// TIA Portal project "HEAT-1-CADIZ-V24" (V20) (continued)

       CASE #modeRequest OF
           1: // ======= Conceder control a KukaControl =========
               // Requisito: que el otro lado (Supervisor) esté ocioso (Queda por ajustar)
               IF #safeAllOk AND (NOT #autoBusy) THEN

                   // 1) Fijar modo efectivo → AutoExtSeq cargará PGNO = 1
                   #modeEffective := USINT#1;

                   // 2) Aún no estamos listos hasta que AutoExtSeq termine
                   "PlcStatus".mode.ready := FALSE;

                   // 3) Señal PNIO al robot para que salga del bucle autoloop.src (CASE 1 del cell.src)
                   #enterCellCase1 := TRUE;

                   // 4) Arranque de AutoExt: PULSO 1-scan a %M770.0
                   #startAutoExt := TRUE;

                   // 5) Handshake a la HMI con el MISMO seq que se recibió
                   "PlcStatus".exec.ackSeq := #modeReqSeq;
                   "PlcStatus".exec.accepted := TRUE;  // 1 scan
                   "PlcStatus".exec.done := TRUE;  // 1 scan
               END_IF;

           2: // ======= Conceder control a Supervisor/VisualScan =========
               // Requisito: que KukaControl esté ocioso
               IF #safeAllOk AND (NOT #servBusy) THEN

                   // 1) Fijar modo efectivo → AutoExtSeq cargará PGNO = 2
                   #modeEffective := USINT#2;

                   // 2) Aún no estamos listos hasta que AutoExtSeq termine
                   "PlcStatus".mode.ready := FALSE;

                   // 3) Señal PNIO al robot para que salga del bucle actual autoloopsup.src (CASE 2 del cell.src)
                   #enterCellCase2 := TRUE;

                   // 4) Arranque de AutoExt: PULSO 1-scan a %M770.0
                   #startAutoExt := TRUE;

                   // 5) Handshake a la HMI
                   "PlcStatus".exec.ackSeq := #modeReqSeq;
                   "PlcStatus".exec.accepted := TRUE;
                   "PlcStatus".exec.done := TRUE;
               END_IF;
       END_CASE;

   END_IF;
END_REGION
END_FUNCTION_BLOCK

FUNCTION_BLOCK "KukaControlSeq"   // FB21, LAD
{ S7_Optimized_Access := 'TRUE' }
VERSION : 0.1
   VAR
      rEnterAuto : R_TRIG;
   END_VAR
   VAR_TEMP
      _clear990 : Bool;
   END_VAR
BEGIN

REGION Network 2: Envia posiciones a la aplicacion KukaControl
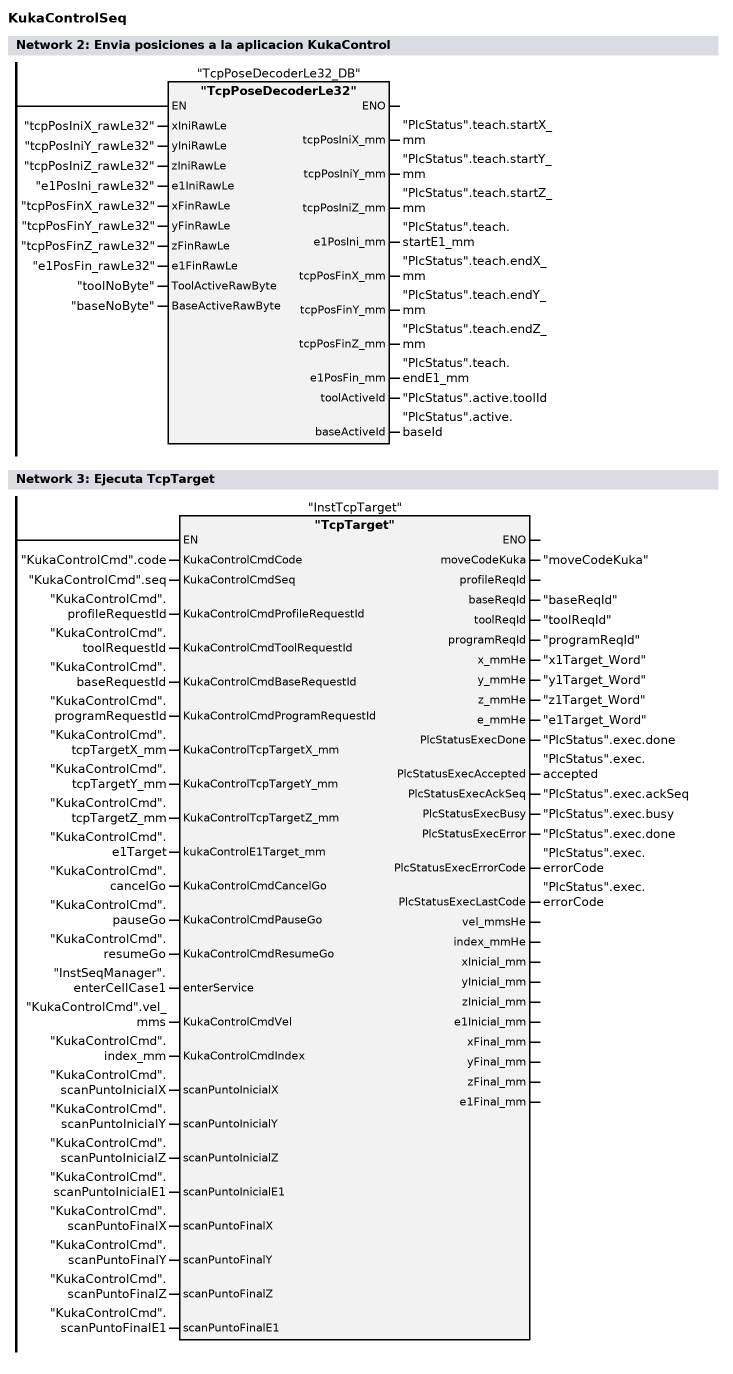
   RUNG wire#powerrail
      "TcpPoseDecoderLe32_DB"(xIniRawLe := "tcpPosIniX_rawLe32", yIniRawLe := "tcpPosIniY_rawLe32", zIniRawLe := "tcpPosIniZ_rawLe32", e1IniRawLe := "e1PosIni_rawLe32", xFinRawLe := "tcpPosFinX_rawLe32", yFinRawLe := "tcpPosFinY_rawLe32", zFinRawLe := "tcpPosFinZ_rawLe32", e1FinRawLe := "e1PosFin_rawLe32", ToolActiveRawByte := "toolNoByte", BaseActiveRawByte := "baseNoByte", tcpPosIniX_mm => "PlcStatus".teach.startX_mm, tcpPosIniY_mm => "PlcStatus".teach.startY_mm, tcpPosIniZ_mm => "PlcStatus".teach.startZ_mm, e1PosIni_mm => "PlcStatus".teach.startE1_mm, tcpPosFinX_mm => "PlcStatus".teach.endX_mm, tcpPosFinY_mm => "PlcStatus".teach.endY_mm, tcpPosFinZ_mm => "PlcStatus".teach.endZ_mm, e1PosFin_mm => "PlcStatus".teach.endE1_mm, toolActiveId => "PlcStatus".active.toolId, baseActiveId => "PlcStatus".active.baseId)
   END_RUNG
   // the same network as SCL:
   "TcpPoseDecoderLe32_DB"(xIniRawLe := "tcpPosIniX_rawLe32",   // "TcpPoseDecoderLe32"
                           yIniRawLe := "tcpPosIniY_rawLe32",
                           zIniRawLe := "tcpPosIniZ_rawLe32",
                           e1IniRawLe := "e1PosIni_rawLe32",
                           xFinRawLe := "tcpPosFinX_rawLe32",
                           yFinRawLe := "tcpPosFinY_rawLe32",
                           zFinRawLe := "tcpPosFinZ_rawLe32",
                           e1FinRawLe := "e1PosFin_rawLe32",
                           ToolActiveRawByte := "toolNoByte",
                           BaseActiveRawByte := "baseNoByte",
                           tcpPosIniX_mm => "PlcStatus".teach.startX_mm,
                           tcpPosIniY_mm => "PlcStatus".teach.startY_mm,
                           tcpPosIniZ_mm => "PlcStatus".teach.startZ_mm,
                           e1PosIni_mm => "PlcStatus".teach.startE1_mm,
                           tcpPosFinX_mm => "PlcStatus".teach.endX_mm,
                           tcpPosFinY_mm => "PlcStatus".teach.endY_mm,
                           tcpPosFinZ_mm => "PlcStatus".teach.endZ_mm,
                           e1PosFin_mm => "PlcStatus".teach.endE1_mm,
                           toolActiveId => "PlcStatus".active.toolId,
                           baseActiveId => "PlcStatus".active.baseId);
END_REGION

REGION Network 3: Ejecuta TcpTarget
   RUNG wire#powerrail
      "InstTcpTarget"(KukaControlCmdCode := "KukaControlCmd".code, KukaControlCmdSeq := "KukaControlCmd".seq, KukaControlCmdProfileRequestId := "KukaControlCmd".profileRequestId, KukaControlCmdToolRequestId := "KukaControlCmd".toolRequestId, KukaControlCmdBaseRequestId := "KukaControlCmd".baseRequestId, KukaControlCmdProgramRequestId := "KukaControlCmd".programRequestId, KukaControlTcpTargetX_mm := "KukaControlCmd".tcpTargetX_mm, KukaControlTcpTargetY_mm := "KukaControlCmd".tcpTargetY_mm, KukaControlTcpTargetZ_mm := "KukaControlCmd".tcpTargetZ_mm, kukaControlE1Target_mm := "KukaControlCmd".e1Target, KukaControlCmdCancelGo := "KukaControlCmd".cancelGo, KukaControlCmdPauseGo := "KukaControlCmd".pauseGo, KukaControlCmdResumeGo := "KukaControlCmd".resumeGo, enterService := "InstSeqManager".enterCellCase1, KukaControlCmdVel := "KukaControlCmd".vel_mms, KukaControlCmdIndex := "KukaControlCmd".index_mm, scanPuntoInicialX := "KukaControlCmd".scanPuntoInicialX, scanPuntoInicialY := "KukaControlCmd".scanPuntoInicialY, scanPuntoInicialZ := "KukaControlCmd".scanPuntoInicialZ, scanPuntoInicialE1 := "KukaControlCmd".scanPuntoInicialE1, scanPuntoFinalX := "KukaControlCmd".scanPuntoFinalX, scanPuntoFinalY := "KukaControlCmd".scanPuntoFinalY, scanPuntoFinalZ := "KukaControlCmd".scanPuntoFinalZ, scanPuntoFinalE1 := "KukaControlCmd".scanPuntoFinalE1, moveCodeKuka => "moveCodeKuka", profileReqId =>, baseReqId => "baseReqId", toolReqId => "toolReqId", programReqId => "programReqId", x_mmHe => "x1Target_Word", y_mmHe => "y1Target_Word", z_mmHe => "z1Target_Word", e_mmHe => "e1Target_Word", PlcStatusExecDone => "PlcStatus".exec.done, PlcStatusExecAccepted => "PlcStatus".exec.accepted, PlcStatusExecAckSeq => "PlcStatus".exec.ackSeq, PlcStatusExecBusy => "PlcStatus".exec.busy, PlcStatusExecError => "PlcStatus".exec.done, PlcStatusExecErrorCode => "PlcStatus".exec.errorCode, PlcStatusExecLastCode => "PlcStatus".exec.errorCode, vel_mmsHe =>, index_mmHe =>, xInicial_mm =>, yInicial_mm =>, zInicial_mm =>, e1Inicial_mm =>, xFinal_mm =>, yFinal_mm =>, zFinal_mm =>, e1Final_mm =>)
   END_RUNG
   // the same network as SCL:
   "InstTcpTarget"(KukaControlCmdCode := "KukaControlCmd".code,   // "TcpTarget"
                   KukaControlCmdSeq := "KukaControlCmd".seq,
                   KukaControlCmdProfileRequestId := "KukaControlCmd".profileRequestId,
                   KukaControlCmdToolRequestId := "KukaControlCmd".toolRequestId,
                   KukaControlCmdBaseRequestId := "KukaControlCmd".baseRequestId,
                   KukaControlCmdProgramRequestId := "KukaControlCmd".programRequestId,
                   KukaControlTcpTargetX_mm := "KukaControlCmd".tcpTargetX_mm,
                   KukaControlTcpTargetY_mm := "KukaControlCmd".tcpTargetY_mm,
                   KukaControlTcpTargetZ_mm := "KukaControlCmd".tcpTargetZ_mm,
                   kukaControlE1Target_mm := "KukaControlCmd".e1Target,
                   KukaControlCmdCancelGo := "KukaControlCmd".cancelGo,
                   KukaControlCmdPauseGo := "KukaControlCmd".pauseGo,
                   KukaControlCmdResumeGo := "KukaControlCmd".resumeGo,
                   enterService := "InstSeqManager".enterCellCase1,
                   KukaControlCmdVel := "KukaControlCmd".vel_mms,
                   KukaControlCmdIndex := "KukaControlCmd".index_mm,
                   scanPuntoInicialX := "KukaControlCmd".scanPuntoInicialX,
                   scanPuntoInicialY := "KukaControlCmd".scanPuntoInicialY,
                   scanPuntoInicialZ := "KukaControlCmd".scanPuntoInicialZ,
                   scanPuntoInicialE1 := "KukaControlCmd".scanPuntoInicialE1,
                   scanPuntoFinalX := "KukaControlCmd".scanPuntoFinalX,
                   scanPuntoFinalY := "KukaControlCmd".scanPuntoFinalY,
                   scanPuntoFinalZ := "KukaControlCmd".scanPuntoFinalZ,
                   scanPuntoFinalE1 := "KukaControlCmd".scanPuntoFinalE1,
                   moveCodeKuka => "moveCodeKuka",
                   baseReqId => "baseReqId",
                   toolReqId => "toolReqId",
                   programReqId => "programReqId",
                   x_mmHe => "x1Target_Word",
                   y_mmHe => "y1Target_Word",
                   z_mmHe => "z1Target_Word",
                   e_mmHe => "e1Target_Word",
                   PlcStatusExecDone => "PlcStatus".exec.done,
                   PlcStatusExecAccepted => "PlcStatus".exec.accepted,
                   PlcStatusExecAckSeq => "PlcStatus".exec.ackSeq,
                   PlcStatusExecBusy => "PlcStatus".exec.busy,
                   PlcStatusExecError => "PlcStatus".exec.done,
                   PlcStatusExecErrorCode => "PlcStatus".exec.errorCode,
                   PlcStatusExecLastCode => "PlcStatus".exec.errorCode);
END_REGION

REGION Network 4 (SCL)
   IF #_clear990 THEN
       "KukaControlCmd".code := 0;                     // no “ensucia” el DB
       #_clear990 := FALSE;
   END_IF;
END_REGION
END_FUNCTION_BLOCK

FUNCTION_BLOCK "SupervisorSeq"   // FB22, LAD
{ S7_Optimized_Access := 'TRUE' }
VERSION : 0.1
   VAR_INPUT
      T_Heartbeat : Time := T#1000ms;   // Periodo del heartbeat PLC
      T_IdCheck : Time := T#2000ms;   // Duración simulada de Identification (comprobaciones)
      enable : Bool;   // Habilita FB -> PLC.plc_ok
      QR_Ready : Bool := true;   // Hay un ID de carrito leído
      CarriageID : String := 'null';   // ID de carrito leído por QR
      TeachAtStart : Bool;   // Teaching (pág. 4): robot en punto de inicio de la siguiente trayectoria
      kukaAtPerspexPos : Bool;   // PA check (Perspex) y Balancing (pág. 6): Robot posicionado en Perspex
      kukaAtGainPos : Bool;   // Gain (pág. 7) -Robot posicionado para Gain
      kukaAtTCGPos : Bool;   // TCG (pág. 8) — multiposición Robot en la posición TCG actual
      kukaAtRefScanStartPos : Bool;   // Robot listo para Scan Ref
      kukaAtInspScanStartPos : Bool;   // Robot listo para Scan Insp
      kukaRefScanFinished : Bool;   // Trayectoria de referencia terminada (robot/UT)
      kukaInspScanFinished : Bool;   // Trayectoria de inspección terminada (robot/UT)
      StartUSReady : Bool := TRUE;   // StartUS (pág. 5): end-effector y precondiciones listas -- True cuando “previous task done”
      MarkingDone : Bool;   // Pre-eval / marcado (pág. 13) -Resultado del marcado (true=OK)
      CmdStopUS : Bool;   // Orden local para Stop US
      CmdBreakUS : Bool;   // Pulso local Break US
      CmdUnbreakUS : Bool;   // Pulso local Unbreak US
   END_VAR
   VAR_OUTPUT
      ActiveStep : Int;   // Espejo local de PLC.step_plc
      AckSourceDbg : Int;   // Código de fuente de ACK (debug local)
      TCG_NextPosReq : Bool;   // PULSO 1 ciclo: mover a la SIGUIENTE posición TCG
      programReqId : Word;
      moveCodeKuka : Word;
      TCG_AdjustMode : Bool;   // LATCH: TRUE mientras estamos en “ajuste TCG”
   END_VAR
   VAR
      tHeartbeat : TON_TIME;
      hbGate : Bool;
      prevStep : Int := -32768;
      firstScan : Bool;
      teachWasRunning : Bool;
      startUSWasRunning : Bool;
      elemWasRunning : Bool;
      balWasRunning : Bool;
      gainWasRunning : Bool;
      scanRefWasRunning : Bool;
      scanInspWasRunning : Bool;
      L_IdEvalDone : Bool;   // // Identification: ya evalué reqId
      L_tcgNext : Bool;
      L_reqRef : Bool;
      L_reqStop : Bool;
      L_reqTcgAdj : Bool;
      L_reqVerif : Bool;
      L_reqPreEval : Bool;
      L_reqIdent : Bool;
      L_reqMark : Bool;
      carriageLatched : Bool;
      validScanParams : Bool;
      waitingNextTCGPos : Bool;
      Cfg_EndEffector : Int;
      Cfg_TeachReq : Bool;
      Cfg_PaCheckReq : Bool;
      Cfg_TcgReq : Bool;
      Cfg_RefName : String;
      PartProgIdx : UInt := 1;   // // index de programa INSP (pieza)
      RefProgIdx : UInt := 1;   // // index de programa REF (pieza)
      tcgIndex : UInt := 1;   // // posición TCG actual
      WantCode : UInt;
      WantProgId : UInt;
      WantToolId : UInt;
      WantIndex : UInt;
      state : Int;
      lastSeq : UInt;
      SupervisorCmdSeq : UInt;
   END_VAR
   VAR_TEMP
      _clear990 : Bool;
      code_int : UInt;
   END_VAR
   VAR CONSTANT
      cSTEP_ID : Int := 1;   // // Pasos (según resumen del PDF, pág. 1)
      cSTEP_TEACH : Int := 2;
      cSTEP_STARTUS : Int := 3;
      cSTEP_PA_BAL : Int := 4;
      cSTEP_GAIN : Int := 5;
      cSTEP_TCG : Int := 6;
      cSTEP_SCAN_REF : Int := 7;
      cSTEP_SCAN_INSP : Int := 8;
      cSTEP_SCAN_REF_VERIF : Int := 9;
      cSTEP_PRE_EVAL : Int := 10;
      cKUKA_REQ_TOOL : UInt := 201;
      cKUKA_GOTO_PERSPEX : UInt := 412;   // mover a Perspex (usa punto enseñado en KRC)
      cKUKA_GOTO_GAIN : UInt := 413;   // mover a Gain
      cKUKA_GOTO_TCG : UInt := 414;   // mover a posición TCG (ARG = index)
      cKUKA_GOTO_REF_START : UInt := 420;   // mover a inicio de Ref (ARG = RefProgIdx)
      cKUKA_GOTO_INSP_START : UInt := 421;   // mover a inicio de Insp (ARG = PartProgIdx)
      cKUKA_RUN_REF_PATH : UInt := 432;   // ejecutar trayectoria de Ref (ARG = RefProgIdx)
      cKUKA_RUN_INSP_PATH : UInt := 433;   // ejecutar trayectoria de Insp (ARG = PartProgIdx)
   END_VAR
BEGIN

REGION Network 1 (SCL)
   // ------------------------------------------------------------------
   // 0) Servicios globales (Heartbeat, housekeeping) — vars generales (pág. 2)
   // ------------------------------------------------------------------
   "PlcStatus".plcOk := #enable;         // espejo de habilitación

   // Heartbeat PLC: toggle con TON (patrón de "compuerta")
   // hbGate se pone TRUE -> TON corre hasta PT -> tHeartbeat.Q = TRUE -> togglamos
   // y bajamos hbGate para reiniciar el ciclo.
   #tHeartbeat(IN := #hbGate,
               PT := #T_Heartbeat);
   IF NOT #hbGate THEN
       #hbGate := TRUE;
   ELSIF #tHeartbeat.Q THEN
       "PlcStatus".heartbeatPlc := NOT "PlcStatus".heartbeatPlc;
       #hbGate := FALSE;
   END_IF;

   // Normalizar paso y espejarlo a salida
   IF ("PlcStatus".stepPlc < #cSTEP_ID) OR ("PlcStatus".stepPlc > #cSTEP_PRE_EVAL) THEN
       "PlcStatus".stepPlc := #cSTEP_ID;
   END_IF;
   #ActiveStep := "PlcStatus".stepPlc;

   // firstScan: 1 ciclo al entrar en cada paso -> útil para resets seguros
   #firstScan := ("PlcStatus".stepPlc <> #prevStep);
   IF #firstScan THEN
       // Limpiamos cualquier "ready/start" que no deba arrastrarse al paso nuevo
       "PlcStatus".startUsReady := FALSE;
       "PlcStatus".stopUsReady := FALSE;
       "PlcStatus".paCheckReady := FALSE;
       "PlcStatus".gainReady := FALSE;
       "PlcStatus".tcgReady := FALSE;
       "PlcStatus".scanRefStart := FALSE;
       "PlcStatus".scanInspStart := FALSE;
       "PlcStatus".markRunning := FALSE;

       // Latches de “estaba corriendo”
       #teachWasRunning := FALSE;
       #startUSWasRunning := FALSE;
       #elemWasRunning := FALSE;
       #balWasRunning := FALSE;
       #gainWasRunning := FALSE;
       #scanRefWasRunning := FALSE;
       #scanInspWasRunning := FALSE;

       // Latches de peticiones (se “arman” al estado actual para evitar disparos al entrar)
       #L_tcgNext := "SupervisorCmd".tcgNextStep;
       #L_reqRef := "SupervisorCmd".reqRefPart;
       #L_reqStop := "SupervisorCmd".reqStopCycle;
       #L_reqTcgAdj := "SupervisorCmd".reqTcgAdj;
       #L_reqVerif := "SupervisorCmd".reqVerif;
       #L_reqPreEval := "SupervisorCmd".reqPreEval;
       #L_reqIdent := "SupervisorCmd".reqIdentificationState;
       #L_reqMark := "SupervisorCmd".reqMark;

       // Identification
       "PlcStatus".idRunning := FALSE;
       #L_IdEvalDone := FALSE;

       // TCG
       #waitingNextTCGPos := ("PlcStatus".stepPlc = #cSTEP_TCG) AND (NOT #kukaAtTCGPos);
       IF "PlcStatus".stepPlc <> #cSTEP_TCG THEN
           #tcgIndex := 1;
       END_IF;

       // Vaciar slot de orden pendiente a robot
       #WantCode := 0;
       #WantProgId := 0;
       #WantToolId := 0;
       #WantIndex := 0;

       #prevStep := "PlcStatus".stepPlc;
   END_IF;

   // ------------------------------------------------------------------
   //[1] MÁQUINA DE ESTADOS (OPC UA + disparos al KUKA por goTrigger)
   // ------------------------------------------------------------------
   CASE "PlcStatus".stepPlc OF

           // ===============================================================
           // 1) IDENTIFICATION (pág. 3)
           // ===============================================================
       #cSTEP_ID:
           // --- Handshake de carriage ID ---
           // FÍSICO: lectura real de QR/PNs/params en KukaControl.
           // El PLC refleja ID leído y valida condiciones base (safety, agua, robot OK).
           // Supervisor.req_carriage_id = TRUE -> el PLC debe mandar:
           //   PLC.carriage_Id (string) y PLC.new_carriage_Id = TRUE
           // Mientras dure la petición. Al bajar la petición, el PLC
           // limpia new_carriage_Id y deja de enviar.
           // req_carriage_id: enviar ID nuevo UNA VEZ mientras Supervisor lo solicite
           IF "SupervisorCmd".reqCarriageId THEN
               IF #QR_Ready AND NOT #carriageLatched  THEN
                   #CarriageID := 'Id de Prueba';
                   "PlcStatus".carriageId := #CarriageID; // escribimos el ID leído
                   "PlcStatus".newCarriageId := TRUE;     // “ID listo”
                   #carriageLatched  := TRUE;              // evita rearmar en el mismo pulso
               END_IF;
           ELSE
               // fin del handshake
               "PlcStatus".newCarriageId := FALSE;
               #carriageLatched  := FALSE;
           END_IF;

           // --- req_id (latch: eval una sola vez en “alto” y decidir salto al bajar) ---
           "PlcStatus".idRunning := "SupervisorCmd".reqId;

           // 1) Primera vez con reqId=TRUE → congelar configuración + calcular id_ok
           IF "SupervisorCmd".reqId AND NOT #L_IdEvalDone THEN
               // Congelar lo que Supervisor ha decidido para el ciclo
               #Cfg_EndEffector := "SupervisorCmd".endEffector;  // 1..5
               #Cfg_TeachReq := "SupervisorCmd".teachReq;
               #Cfg_PaCheckReq := "SupervisorCmd".paCheckReq;
               #Cfg_TcgReq := "SupervisorCmd".tcgReq;
               #Cfg_RefName := "SupervisorCmd".referencePart;

               // Resolver índices de programa por pieza
               // >>> AJUSTAR a los nombres reales de piezas/referencias <<<
               IF #Cfg_RefName = 'PIEZA1' THEN
                   #PartProgIdx := 1;
                   #RefProgIdx := 1;
               ELSIF #Cfg_RefName = 'PIEZA2' THEN
                   #PartProgIdx := 2;
                   #RefProgIdx := 2;
               ELSIF #Cfg_RefName = 'PIEZA3' THEN
                   #PartProgIdx := 3;
                   #RefProgIdx := 3;
               ELSE
                   #PartProgIdx := 1;
                   #RefProgIdx := 1;
               END_IF;

               // id_ok = enclavamientos + servicios + herramienta válida
               "PlcStatus".idOk :=
               ("PlcStatus".plcOk AND "SupervisorCmd".supervisorOk AND "PlcStatus".robotOk AND "PlcStatus".safetyOk
               AND "PlcStatus".airOk AND "PlcStatus".inspWaterOk AND "PlcStatus".tankWaterOk)
               AND (#Cfg_EndEffector >= 1) AND (#Cfg_EndEffector <= 5);

               #L_IdEvalDone := TRUE; // evita re‑evaluar cada scan mientras reqId siga alto
           END_IF;

           // 2) Cuando reqId cae a FALSE → decidir próximo paso
           IF (NOT "SupervisorCmd".reqId) AND #L_IdEvalDone THEN
               IF NOT "PlcStatus".idOk THEN
                   "PlcStatus".stepPlc := #cSTEP_ID;          // quedarse en Identification
               ELSE
                   IF #Cfg_TeachReq THEN
                       "PlcStatus".stepPlc := #cSTEP_TEACH;   // ir a Teaching
                   ELSE
                       "PlcStatus".stepPlc := #cSTEP_STARTUS; // ir a inicio UT
                   END_IF;
               END_IF;
               #L_IdEvalDone := FALSE; // rearmado para la próxima identificación
           END_IF;


           // ===============================================================
           // 2) TEACHING (pág. 4) — multi-PN: rearmar teach_ready por PN
           // FÍSICO: si la herramienta necesaria para teaching no está montada,
           // el KUKA cambia en Staübli al stand indicado (usa Supervisor.end-effector).
           // Luego, el KUKA se mueve al INICIO del PN siguiente y pone un bit de “en posición”.
           // Ese bit alimenta TeachAtStart=TRUE. Entonces EL PLC arma teach_ready (p. 4).
           // Repetir por cada PN mientras teach_app_running=TRUE.
           // ===============================================================
           (*  #cSTEP_TEACH:

             IF "SupervisorCmd".teachAppRunning THEN
                   IF (NOT "SupervisorCmd".teachRunning) AND TeachAtStart THEN
                       "PlcStatus".teachReady := TRUE;
                   END_IF;

                   IF "SupervisorCmd".teachRunning THEN
                       "PlcStatus".teachReady := FALSE;
                       teachWasRunning := TRUE;
                   END_IF;

                   // Fin de una trayectoria de teaching (sin abandonar la app)
                   IF (NOT "SupervisorCmd".teachRunning) AND teachWasRunning THEN
                       teachWasRunning := FALSE;
                   END_IF;

               ELSE
                   // Cierre de la app: salto según teach_state
                   IF "SupervisorCmd".teachState THEN
                       "PlcStatus".stepPlc := cSTEP_STARTUS;
                   ELSE
                       "PlcStatus".stepPlc := cSTEP_ID;
                   END_IF;
               END_IF;
           END_IF;*)




           // ===============================================================
           // 3) START US (pág. 5) — armar cuando “previous task done”
           // FÍSICO: KUKA AUT EXT cambia (si hace falta) al efector de INSPECCIÓN
           // requerido (Supervisor.end-effector, p. 1). Cuando:
           //   - Herramienta correcta acoplada (Staübli OK),
           //   - servicios/enclavamientos OK (safety/air/water/tank),
           //   - robot en posición segura para inicializar el UT,
           // el secuenciador pone StartUSReady=TRUE. El PLC arma start_us_ready.
           // Supervisor hace init UT (start_us_running/state_us). (p. 5)
           // ===============================================================
       #cSTEP_STARTUS:

           // Al entrar, ordena al robot cargar la herramienta decidida en ID
           IF #firstScan THEN
               #SupervisorCmdSeq := #SupervisorCmdSeq + 1;
               #WantCode := #cKUKA_REQ_TOOL;
               #WantToolId := (#Cfg_EndEffector);       // 1..5
           END_IF;

           // El PLC arma startUsReady SI el entorno/robot están listos y todavía no corre
           IF #StartUSReady AND NOT "SupervisorCmd".startUsRunning THEN
               "PlcStatus".startUsReady := TRUE;
           END_IF;

           // Cuando arranca, baja el "ready" y registra que realmente empezó
           IF "SupervisorCmd".startUsRunning THEN
               "PlcStatus".startUsReady := FALSE;
               #startUSWasRunning := TRUE;
           END_IF;

           // Al terminar: salto a PA o a Gain según lo congelado en ID
           IF (NOT "SupervisorCmd".startUsRunning) AND #startUSWasRunning THEN
               #startUSWasRunning := FALSE;
               IF NOT "SupervisorCmd".stateUs THEN
                   "PlcStatus".stepPlc := #cSTEP_ID;
               ELSE
                   IF #Cfg_PaCheckReq THEN
                       "PlcStatus".stepPlc := #cSTEP_PA_BAL;
                   ELSE
                       "PlcStatus".stepPlc := #cSTEP_GAIN;
                   END_IF;
               END_IF;
           END_IF;


           // ===============================================================
           // 4) DEAD ELEMENT CHECK & BALANCING (pág. 6)
           //FÍSICO: KUKA va a la pieza Perspex de calibración y, cuando está en
           // posición estática, tu lógica pone AtPerspex=TRUE. El PLC arma
           // pa_check_ready y el Supervisor ejecuta elem_running/bal_running (p. 6).
           // ===============================================================
       #cSTEP_PA_BAL:

           // Posicionamiento automático a Perspex si no estamos ya
           IF (NOT #kukaAtPerspexPos) AND (#WantCode = 0) THEN
               #SupervisorCmdSeq := #SupervisorCmdSeq + 1;
               #WantCode := #cKUKA_GOTO_PERSPEX;
           END_IF;

           // Armado del ready cuando estemos en Perspex y aún no corre elem_running
           IF #kukaAtPerspexPos AND NOT "SupervisorCmd".elemRunning THEN
               "PlcStatus".paCheckReady := TRUE;
           END_IF;

           IF "SupervisorCmd".elemRunning THEN
               "PlcStatus".paCheckReady := FALSE;
               #elemWasRunning := TRUE;
           END_IF;

           IF (NOT "SupervisorCmd".elemRunning) AND #elemWasRunning THEN
               #elemWasRunning := FALSE;
               IF NOT "SupervisorCmd".elemState THEN
                   "PlcStatus".stepPlc := #cSTEP_ID;
               ELSE
                   // Encadenar balancing (igual patrón running/state)
                   IF "SupervisorCmd".balRunning THEN
                       #balWasRunning := TRUE;
                   END_IF;

                   IF (NOT "SupervisorCmd".balRunning) AND #balWasRunning THEN
                       #balWasRunning := FALSE;
                       IF "SupervisorCmd".balState THEN
                           "PlcStatus".stepPlc := #cSTEP_GAIN;
                       ELSE
                           "PlcStatus".stepPlc := #cSTEP_ID;
                       END_IF;
                   END_IF;
               END_IF;
           END_IF;

           // ===============================================================
           // 5) GAIN ADJUSTMENT (pág. 7)
           // FÍSICO: KUKA se posiciona en la referencia para ganancia estática;
           // cuando está “en posición”, AtGainPos=TRUE. PLC arma gain_ready;
           // Supervisor ejecuta gain_running/gain_state y decide si ir a TCG (p. 7).
           // ===============================================================
       #cSTEP_GAIN:

           // Posicionamiento a Gain si no estamos ya
           IF (NOT #kukaAtGainPos) AND (#WantCode = 0) THEN
               #SupervisorCmdSeq := #SupervisorCmdSeq + 1;
               #WantCode := #cKUKA_GOTO_GAIN;
           END_IF;

           IF #kukaAtGainPos AND NOT "SupervisorCmd".gainRunning THEN
               "PlcStatus".gainReady := TRUE;
           END_IF;

           IF "SupervisorCmd".gainRunning THEN
               "PlcStatus".gainReady := FALSE;
               #gainWasRunning := TRUE;
           END_IF;

           IF (NOT "SupervisorCmd".gainRunning) AND #gainWasRunning THEN
               #gainWasRunning := FALSE;
               IF NOT "SupervisorCmd".gainState THEN
                   "PlcStatus".stepPlc := #cSTEP_ID;
               ELSE
                   IF #Cfg_TcgReq THEN
                       "PlcStatus".stepPlc := #cSTEP_TCG;
                   ELSE
                       "PlcStatus".stepPlc := #cSTEP_SCAN_REF;
                   END_IF;
               END_IF;
           END_IF;

           // ===============================================================
           // (6) TCG CHECK / ADJUSTMENT — pág. 8 (multiposición)
           // FÍSICO: KUKA recorre varias posiciones TCG. Para cada posición:
           //   - Cuando el robot está en la POSICIÓN TCG ACTUAL (estático),
           //     tu lógica pone AtTCGPos=TRUE → PLC arma tcg_ready (p. 8).
           //   - Supervisor pone tcg_in_progress=TRUE mientras mide.
           //   - Al pulsar “Next” en Supervisor (tcg_next_step=TRUE), el ACK manager
           //     emite TCG_NextPosReq (pulso) para que MUEVAS el robot a la SIGUIENTE
           //     posición; el FB bloquea el rearme (waitingNextTCGPos=TRUE) hasta que
           //     AtTCGPos vuelva a TRUE en la nueva posición (antirrebote).
           //   - Final: según req_ref_part / req_stop_cycle / req_tcg_adj (p. 8).
           // ===============================================================
       #cSTEP_TCG:

           // Si acabamos de entrar y no estamos en la pos TCG actual, pedir el movimiento
           IF (NOT #kukaAtTCGPos) AND (#WantCode = 0) AND (NOT #waitingNextTCGPos) THEN
               #SupervisorCmdSeq := #SupervisorCmdSeq + 1;
               #WantCode := #cKUKA_GOTO_TCG;
               #WantIndex := (#tcgIndex);     // índice a mover
               #waitingNextTCGPos := TRUE;
           END_IF;

           // Rearme de espera cuando lleguemos
           IF #waitingNextTCGPos AND #kukaAtTCGPos THEN
               #waitingNextTCGPos := FALSE;
           END_IF;

           // tcg_ready sólo si no mide y no esperamos pos
           IF (NOT "SupervisorCmd".tcgInProgress) AND (NOT #waitingNextTCGPos) THEN
               "PlcStatus".tcgReady := TRUE;
           END_IF;

           IF "SupervisorCmd".tcgInProgress THEN
               "PlcStatus".tcgReady := FALSE;
           END_IF;

           // NEXT (una vez por pulsación): incrementar índice y ordenar movimiento
           IF "SupervisorCmd".tcgNextStep AND NOT #L_tcgNext THEN
               #SupervisorCmdSeq := #SupervisorCmdSeq + 1;
               #tcgIndex := #tcgIndex + 1;
               #WantCode := #cKUKA_GOTO_TCG;
               #WantIndex := (#tcgIndex);
               #waitingNextTCGPos := TRUE;
               #L_tcgNext := TRUE;
           END_IF;
           IF NOT "SupervisorCmd".tcgNextStep THEN
               #L_tcgNext := FALSE;
           END_IF;

           // Decisiones finales (una sola vez)
           IF "SupervisorCmd".reqRefPart AND NOT #L_reqRef THEN
               "PlcStatus".stepPlc := #cSTEP_SCAN_REF;
               #L_reqRef := TRUE;
           END_IF;
           IF NOT "SupervisorCmd".reqRefPart THEN
               #L_reqRef := FALSE;
           END_IF;

           IF "SupervisorCmd".reqStopCycle AND NOT #L_reqStop THEN
               "PlcStatus".stepPlc := #cSTEP_ID;
               #L_reqStop := TRUE;
           END_IF;
           IF NOT "SupervisorCmd".reqStopCycle THEN
               #L_reqStop := FALSE;
           END_IF;

           IF "SupervisorCmd".reqTcgAdj AND NOT #L_reqTcgAdj THEN
               // permanecer en TCG en modo ajuste (no cambia de paso)
               #L_reqTcgAdj := TRUE;
           END_IF;
           IF NOT "SupervisorCmd".reqTcgAdj THEN
               #L_reqTcgAdj := FALSE;
           END_IF;



           // ===============================================================
           // (7) SCAN REFERENCE ACQUISITION — pág. 10
           // FÍSICO: KUKA carga PN/frame y se coloca en el punto de INICIO de
           // la trayectoria de referencia. Tu lógica pone AtRefScanStart=TRUE cuando
           // está en posición. El PLC solo arma scan_ref_start si además los
           // parámetros mínimos (id_scan, x_size, y_size) están válidos (p. 10).
           // ===============================================================
       #cSTEP_SCAN_REF:

           // Validación mínima de parámetros de scan que el PLC publica al Supervisor
           #validScanParams := (LEN("PlcStatus".idScan) > 0) AND ("PlcStatus".xSize > 0.0) AND ("PlcStatus".ySize > 0.0);

           // Posicionar al inicio de Ref si no estamos (CASE 420, ARG=RefProgIdx)
           IF (NOT #kukaAtRefScanStartPos) AND (#WantCode = 0) THEN
               #SupervisorCmdSeq := #SupervisorCmdSeq + 1;
               #WantCode := #cKUKA_GOTO_REF_START; // ← KRC: CASE 420
               #WantProgId := (#RefProgIdx);   // índice de programa REF por pieza
           END_IF;

           // Permiso de arranque
           IF #kukaAtRefScanStartPos AND #validScanParams AND NOT "SupervisorCmd".scanRefRunning THEN
               "PlcStatus".scanRefStart := TRUE;   // ← Anunciar “ready” al Supervisor
           END_IF;

